
           #statSend.tsendFct.data[#statSend.tsendFct.dataOffset + 8] := #statSend.dataTelegram.ackMessageOffset.%B3;
           #statSend.tsendFct.data[#statSend.tsendFct.dataOffset + 9] := #statSend.dataTelegram.ackMessageOffset.%B2;
           #statSend.tsendFct.data[#statSend.tsendFct.dataOffset + 10] := #statSend.dataTelegram.ackMessageOffset.%B1;
           #statSend.tsendFct.data[#statSend.tsendFct.dataOffset + 11] := #statSend.dataTelegram.ackMessageOffset.%B0;

           #statSend.tsendFct.data[#statSend.tsendFct.dataOffset + 12] := #statSend.dataTelegram.actPackageLength.%B3;
           #statSend.tsendFct.data[#statSend.tsendFct.dataOffset + 13] := #statSend.dataTelegram.actPackageLength.%B2;
           #statSend.tsendFct.data[#statSend.tsendFct.dataOffset + 14] := #statSend.dataTelegram.actPackageLength.%B1;
           #statSend.tsendFct.data[#statSend.tsendFct.dataOffset + 15] := #statSend.dataTelegram.actPackageLength.%B0;

           #statSend.tsendFct.data[#statSend.tsendFct.dataOffset + 16] := #statSend.dataTelegram.totalMessageLength.%B3;
           #statSend.tsendFct.data[#statSend.tsendFct.dataOffset + 17] := #statSend.dataTelegram.totalMessageLength.%B2;
           #statSend.tsendFct.data[#statSend.tsendFct.dataOffset + 18] := #statSend.dataTelegram.totalMessageLength.%B1;
           #statSend.tsendFct.data[#statSend.tsendFct.dataOffset + 19] := #statSend.dataTelegram.totalMessageLength.%B0;

           //LCom V2
           IF (#diagnostics.statistics.activeLComVersion = #LCOM_HEADER_V2) THEN
             //Calculate offset in the tcp send buffer
             #statSend.tsendFct.dataOffset := #statSend.tsendFct.dataOffset + 20;
           ELSE
             //LCom V1
             //MessageOffset
             #statSend.tsendFct.data[#statSend.tsendFct.dataOffset + 4] := #statSend.dataTelegram.messageOffset.%B1;
             #statSend.tsendFct.data[#statSend.tsendFct.dataOffset + 5] := #statSend.dataTelegram.messageOffset.%B0;
             //AckMessageOffset
             #statSend.tsendFct.data[#statSend.tsendFct.dataOffset + 6] := #statSend.dataTelegram.ackMessageOffset.%B1;
             #statSend.tsendFct.data[#statSend.tsendFct.dataOffset + 7] := #statSend.dataTelegram.ackMessageOffset.%B0;
             //ActPackageLength
             #statSend.tsendFct.data[#statSend.tsendFct.dataOffset + 8] := #statSend.dataTelegram.actPackageLength.%B1;
             #statSend.tsendFct.data[#statSend.tsendFct.dataOffset + 9] := #statSend.dataTelegram.actPackageLength.%B0;
             //TotalMessageLength
             #statSend.tsendFct.data[#statSend.tsendFct.dataOffset + 10] := #statSend.dataTelegram.totalMessageLength.%B1;
             #statSend.tsendFct.data[#statSend.tsendFct.dataOffset + 11] := #statSend.dataTelegram.totalMessageLength.%B0;
             //Calculate offset in the tcp send buffer
             #statSend.tsendFct.dataOffset := #statSend.tsendFct.dataOffset + 12;
           END_IF;

           //Store expected acknowledge message offset and time
           #statSend.expectedAck.package1.offset := #statSend.dataTelegram.messageOffset + #statSend.dataTelegram.actPackageLength;
           //Start expe. message Timer 1
           #instExpectedAckPackage1(IN := TRUE,
                                    PT := #diagnostics.localConfig.sender.ackTimeout);

           #statSend.numberOfLComPackage := #statSend.numberOfLComPackage + 1;

           //Copy data from FB.sendBuffer
           #statRet := MOVE_BLK_VARIANT(SRC := #sendBuffer, COUNT := #statSend.dataTelegram.actPackageLength, SRC_INDEX := UDINT_TO_DINT(#statSend.userData.offset), DEST_INDEX := #statSend.tsendFct.dataOffset, DEST => #statSend.tsendFct.data);
           //Calculate offset in FB.sendBuffer
           #statSend.userData.offset := #statSend.userData.offset + #statSend.dataTelegram.actPackageLength;
           //Copy offset in telegram
           #statSend.dataTelegram.messageOffset := #statSend.userData.offset;
           //Calculate offset in the tcp send buffer
           #statSend.tsendFct.dataOffset := #statSend.tsendFct.dataOffset + UDINT_TO_UINT(#statSend.dataTelegram.actPackageLength);

           //All sent data is copied ?
           IF (#statSend.userData.offset = #statSend.dataTelegram.totalMessageLength) THEN
             //Yes
             #statState.comSender := #SEND_NO_DATA;
           ELSE
             ;//No --> Not all sent data has been copied
           END_IF;
         ELSIF (#statState.comSender = #CYCLE
           AND
           (NOT #diagnostics.localConfig.connection.useLComProtocol)) THEN
           //---------------------------------------------------------------------
           //Send telegram without LCom protocol
           //---------------------------------------------------------------------
           #statState.sender := #SEND_DATA;

           //Calculate rest data from the total message
           IF ((#statSend.dataTelegram.totalMessageLength - #statSend.userData.offset) > #MAX_DATA_BUFFER) THEN
             #statSend.tsendFct.dataOffset := #MAX_DATA_BUFFER;
           ELSE
             #statSend.tsendFct.dataOffset := UDINT_TO_UINT(#statSend.dataTelegram.totalMessageLength - #statSend.userData.offset);
           END_IF;

           //Copy data from FB.sendBuffer
           #statRet := MOVE_BLK_VARIANT(SRC := #sendBuffer, COUNT := #statSend.tsendFct.dataOffset, SRC_INDEX := UDINT_TO_DINT(#statSend.userData.offset), DEST_INDEX := 0, DEST => #statSend.tsendFct.data);
           //Calculate offset in tcp send buffer
           #statSend.userData.offset := #statSend.userData.offset + #statSend.tsendFct.dataOffset;
           //End: Send telegram without LCom protocol
         ELSE
           ;//Not in sending process 
         END_IF;//End: Send telegram
       END_IF;//End: Connected


       //---------------------------------------------------------------------
       //State machine sender configuration
       //---------------------------------------------------------------------
       CASE #statState.cfgSender OF

         #OPERATION:
           ;//Sender configuration successful exchange
         #STATE_WAIT:
           ;
         #STATE_INIT:

           #statCompare.sender.cycleTime := #configuration.sender.cycleTime;
           #statCompare.sender.ackTimeOut := #configuration.sender.ackTimeout;

           //LCom Version V1.0
           IF (#statActualLocalLComVersion = #LCOM_HEADER_V1) THEN

             //Check max. cycleTime
             IF (#configuration.sender.cycleTime > T#65535ms) THEN

               #statDiag.bufferIndex := #statDiag.bufferIndex + 1;
               #statDiag.buffer[#statDiag.bufferIndex].additionalValue4 := #configuration.sender.cycleTime;
               #statSend.configTelegramV1.cycleTime := 65535;

               #statDiag.buffer[#statDiag.bufferIndex].status := "LCOM_WARN_SEND_CYCLE_LIMITATION";
               #statDiag.buffer[#statDiag.bufferIndex].subFunctionErrorID := 16#0000;
               #statDiag.buffer[#statDiag.bufferIndex].additionalValue1 := 65535.0;
               #statDiag.buffer[#statDiag.bufferIndex].additionalValue2 := 0.0;
               #statDiag.buffer[#statDiag.bufferIndex].additionalValue3 := 0.0;
             ELSE
               #statSend.configTelegramV1.cycleTime := TIME_TO_UINT(#configuration.sender.cycleTime);
             END_IF;

             //Check max. ackTimeOut
             IF (#configuration.sender.ackTimeout > T#65535ms) THEN

               #statDiag.bufferIndex := #statDiag.bufferIndex + 1;
               #statDiag.buffer[#statDiag.bufferIndex].additionalValue4 := #configuration.sender.ackTimeout;
               #statSend.configTelegramV1.ackTimeOut := 65535;

               #statDiag.buffer[#statDiag.bufferIndex].status := "LCOM_WARN_ACK_TIMEOUT_LIMITATION";
               #statDiag.buffer[#statDiag.bufferIndex].subFunctionErrorID := 16#0000;
               #statDiag.buffer[#statDiag.bufferIndex].additionalValue1 := 65535.0;
               #statDiag.buffer[#statDiag.bufferIndex].additionalValue2 := 0.0;
               #statDiag.buffer[#statDiag.bufferIndex].additionalValue3 := 0.0;
             ELSE
               #statSend.configTelegramV1.ackTimeOut := TIME_TO_UINT(#configuration.sender.ackTimeout);
             END_IF;
           ELSE //LCom Version V2.0
             #statSend.configTelegramV2.cycleTime := #configuration.sender.cycleTime;
             #statSend.configTelegramV2.ackTimeOut := #configuration.sender.ackTimeout;
           END_IF;

           #statState.cfgSender := #SEND_CONFIG;

         #SEND_CONFIG:
           #statState.cfgSender := #STATE_WAIT;

           //LCom Version V1.0
           IF (#statActualLocalLComVersion = #LCOM_HEADER_V1) THEN
             #statSend.tsendFct.data[#statSend.tsendFct.dataOffset] := #statSend.configTelegramV1.LComVersion;
             #statSend.tsendFct.data[#statSend.tsendFct.dataOffset + 1] := 16#02;
             #statSend.tsendFct.data[#statSend.tsendFct.dataOffset + 2] := #statSend.configTelegramV1.comMode;//ComMode
             #statSend.tsendFct.data[#statSend.tsendFct.dataOffset + 3] := #statSend.configTelegramV1.slidingWindow;//SlidingWindow
             //cycleTime
             #statSend.tsendFct.data[#statSend.tsendFct.dataOffset + 4] := #statSend.configTelegramV1.cycleTime.%B1;
             #statSend.tsendFct.data[#statSend.tsendFct.dataOffset + 5] := #statSend.configTelegramV1.cycleTime.%B0;
             //ackTimeOut
             #statSend.tsendFct.data[#statSend.tsendFct.dataOffset + 6] := #statSend.configTelegramV1.ackTimeOut.%B1;
             #statSend.tsendFct.data[#statSend.tsendFct.dataOffset + 7] := #statSend.configTelegramV1.ackTimeOut.%B0;
             //lifeSignCycle
             #statSend.tsendFct.data[#statSend.tsendFct.dataOffset + 8] := #statSend.configTelegramV1.lifeSignCycle.%B1;
             #statSend.tsendFct.data[#statSend.tsendFct.dataOffset + 9] := #statSend.configTelegramV1.lifeSignCycle.%B0;
             //status
             #statSend.tsendFct.data[#statSend.tsendFct.dataOffset + 10] := #statSend.configTelegramV1.status;
             //sendModeSyncTime
             #statSend.tsendFct.data[#statSend.tsendFct.dataOffset + 11] := #statSend.configTelegramV1.sendModeSyncTime;
             //maxSendDataLength
             #statSend.tsendFct.data[#statSend.tsendFct.dataOffset + 12] := #statSend.configTelegramV1.maxSendDataLength.%B1;
             #statSend.tsendFct.data[#statSend.tsendFct.dataOffset + 13] := #statSend.configTelegramV1.maxSendDataLength.%B0;
             //maxReceiveDataLength
             #statSend.tsendFct.data[#statSend.tsendFct.dataOffset + 14] := #statSend.configTelegramV1.maxReceiveDataLength.%B1;
             #statSend.tsendFct.data[#statSend.tsendFct.dataOffset + 15] := #statSend.configTelegramV1.maxReceiveDataLength.%B0;

             #statSend.tsendFct.data[#statSend.tsendFct.dataOffset + 16] := #statSend.configTelegramV1.LComVersion;
             #statSend.tsendFct.data[#statSend.tsendFct.dataOffset + 17] := 16#02;
             #statSend.tsendFct.data[#statSend.tsendFct.dataOffset + 18] := #statSend.configTelegramV1.comMode;//ComMode
             #statSend.tsendFct.data[#statSend.tsendFct.dataOffset + 19] := #statSend.configTelegramV1.slidingWindow;//SlidingWindow
             //cycleTime
             #statSend.tsendFct.data[#statSend.tsendFct.dataOffset + 20] := #statSend.configTelegramV1.cycleTime.%B1;
             #statSend.tsendFct.data[#statSend.tsendFct.dataOffset + 21] := #statSend.configTelegramV1.cycleTime.%B0;
             //ackTimeOut
             #statSend.tsendFct.data[#statSend.tsendFct.dataOffset + 22] := #statSend.configTelegramV1.ackTimeOut.%B1;
             #statSend.tsendFct.data[#statSend.tsendFct.dataOffset + 23] := #statSend.configTelegramV1.ackTimeOut.%B0;
             //lifeSignCycle
             #statSend.tsendFct.data[#statSend.tsendFct.dataOffset + 24] := #statSend.configTelegramV1.lifeSignCycle.%B1;
             #statSend.tsendFct.data[#statSend.tsendFct.dataOffset + 25] := #statSend.configTelegramV1.lifeSignCycle.%B0;
             //status
             #statSend.tsendFct.data[#statSend.tsendFct.dataOffset + 26] := #statSend.configTelegramV1.status;
             //sendModeSyncTime
             #statSend.tsendFct.data[#statSend.tsendFct.dataOffset + 27] := #statSend.configTelegramV1.sendModeSyncTime;
             //maxSendDataLength
             #statSend.tsendFct.data[#statSend.tsendFct.dataOffset + 28] := #statSend.configTelegramV1.maxSendDataLength.%B1;
             #statSend.tsendFct.data[#statSend.tsendFct.dataOffset + 29] := #statSend.configTelegramV1.maxSendDataLength.%B0;
             //maxReceiveDataLength
             #statSend.tsendFct.data[#statSend.tsendFct.dataOffset + 30] := #statSend.configTelegramV1.maxReceiveDataLength.%B1;
             #statSend.tsendFct.data[#statSend.tsendFct.dataOffset + 31] := #statSend.configTelegramV1.maxReceiveDataLength.%B0;
             //calculate new offset
             #statSend.tsendFct.dataOffset := #statSend.tsendFct.dataOffset + 32;
             #statState.sender := #SEND_CONFIG;

             #diagnostics.localConfig.sender.cycleTime := UINT_TO_TIME(#statSend.configTelegramV1.cycleTime);
             #diagnostics.localConfig.sender.ackTimeout := UINT_TO_TIME(#statSend.configTelegramV1.ackTimeOut);
           ELSE
             //LCom Version V2.0
             #statSend.tsendFct.data[#statSend.tsendFct.dataOffset] := #statSend.configTelegramV2.LComVersion;
             #statSend.tsendFct.data[#statSend.tsendFct.dataOffset + 1] := 16#02;
             //status
             #statSend.tsendFct.data[#statSend.tsendFct.dataOffset + 2] := #statSend.configTelegramV2.status;
             //sendModeSyncTime
             #statSend.tsendFct.data[#statSend.tsendFct.dataOffset + 3] := #statSend.configTelegramV2.sendModeSyncTime;
             //lifeSignCycle
             #tempDWord := TIME_TO_DWORD(#statSend.configTelegramV2.lifeSignCycle);
             #statSend.tsendFct.data[#statSend.tsendFct.dataOffset + 4] := #tempDWord.%B3;
             #statSend.tsendFct.data[#statSend.tsendFct.dataOffset + 5] := #tempDWord.%B2;
             #statSend.tsendFct.data[#statSend.tsendFct.dataOffset + 6] := #tempDWord.%B1;
             #statSend.tsendFct.data[#statSend.tsendFct.dataOffset + 7] := #tempDWord.%B0;
             //cycleTime
             #tempDWord := TIME_TO_DWORD(#statSend.configTelegramV2.cycleTime);
             #statSend.tsendFct.data[#statSend.tsendFct.dataOffset + 8] := #tempDWord.%B3;
             #statSend.tsendFct.data[#statSend.tsendFct.dataOffset + 9] := #tempDWord.%B2;
             #statSend.tsendFct.data[#statSend.tsendFct.dataOffset + 10] := #tempDWord.%B1;
             #statSend.tsendFct.data[#statSend.tsendFct.dataOffset + 11] := #tempDWord.%B0;
             //ackTimeOut
             #tempDWord := TIME_TO_DWORD(#statSend.configTelegramV2.ackTimeOut);
             #statSend.tsendFct.data[#statSend.tsendFct.dataOffset + 12] := #tempDWord.%B3;
             #statSend.tsendFct.data[#statSend.tsendFct.dataOffset + 13] := #tempDWord.%B2;
             #statSend.tsendFct.data[#statSend.tsendFct.dataOffset + 14] := #tempDWord.%B1;
             #statSend.tsendFct.data[#statSend.tsendFct.dataOffset + 15] := #tempDWord.%B0;
             //maxSendDataLength
             #statSend.tsendFct.data[#statSend.tsendFct.dataOffset + 16] := #statSend.configTelegramV2.maxSendDataLength.%B3;
             #statSend.tsendFct.data[#statSend.tsendFct.dataOffset + 17] := #statSend.configTelegramV2.maxSendDataLength.%B2;
             #statSend.tsendFct.data[#statSend.tsendFct.dataOffset + 18] := #statSend.configTelegramV2.maxSendDataLength.%B1;
             #statSend.tsendFct.data[#statSend.tsendFct.dataOffset + 19] := #statSend.configTelegramV2.maxSendDataLength.%B0;
             //maxReceiveDataLength
             #statSend.tsendFct.data[#statSend.tsendFct.dataOffset + 20] := #statSend.configTelegramV2.maxReceiveDataLength.%B3;
             #statSend.tsendFct.data[#statSend.tsendFct.dataOffset + 21] := #statSend.configTelegramV2.maxReceiveDataLength.%B2;
             #statSend.tsendFct.data[#statSend.tsendFct.dataOffset + 22] := #statSend.configTelegramV2.maxReceiveDataLength.%B1;
             #statSend.tsendFct.data[#statSend.tsendFct.dataOffset + 23] := #statSend.configTelegramV2.maxReceiveDataLength.%B0;

             //calculate new offset
             #statSend.tsendFct.dataOffset := #statSend.tsendFct.dataOffset + 24;
             #statState.sender := #SEND_CONFIG;

             #diagnostics.localConfig.sender.cycleTime := #statSend.configTelegramV2.cycleTime;
             #diagnostics.localConfig.sender.ackTimeout := #statSend.configTelegramV2.ackTimeOut;

             IF #diagnostics.statistics.activeLComVersion = #LCOM_HEADER_V2 THEN
               #connected := TRUE;
               #diagnostics.statistics.LComProtocolUsed := TRUE;
               #diagnostics.statistics.activeLComVersion := #LCOM_HEADER_V2;
               #statState.cfgSender := #OPERATION;

               //Write diagnostics
               #statDiag.bufferIndex := #statDiag.bufferIndex + 1;
               #statDiag.buffer[#statDiag.bufferIndex].status := "LCOM_STATUS_LCOM_CONNECTED_V2";
               #statDiag.buffer[#statDiag.bufferIndex].subFunctionErrorID := 16#0000;
               #statDiag.buffer[#statDiag.bufferIndex].additionalValue1 := 0.0;
               #statDiag.buffer[#statDiag.bufferIndex].additionalValue2 := 0.0;
               #statDiag.buffer[#statDiag.bufferIndex].additionalValue3 := 0.0;
               #statDiag.buffer[#statDiag.bufferIndex].additionalValue4 := T#0ms;
             END_IF;
           END_IF;

           #statCompare.sender.cycleTime := #configuration.sender.cycleTime;
           #statCompare.sender.ackTimeOut := #configuration.sender.ackTimeout;

         #ERROR_STATE:
           ;
         ELSE
           ;// Statement section ELSE
       END_CASE;


       //No telegram 1,2,5 or 10 to  be sent, therefore check whether life sign tel. must be sent
       IF (#statState.sender = #STATE_INACTIVE
         AND
         (#diagnostics.localConfig.connection.lifeSignCycleTime <> T#0ms)
         AND
         #diagnostics.localConfig.connection.useLComProtocol)
       THEN
         #instLocalLifeSignCycleTimer(IN := TRUE,
                                      PT := #diagnostics.localConfig.connection.lifeSignCycleTime);

         IF (#instLocalLifeSignCycleTimer.Q)
         THEN

           //LCom Version V1.0
           IF (#statActualLocalLComVersion = #LCOM_HEADER_V1) THEN

             //LCom Version V1
             #statSend.tsendFct.data[#statSend.tsendFct.dataOffset] := #statSend.configTelegramV1.LComVersion;
             #statSend.tsendFct.data[#statSend.tsendFct.dataOffset + 1] := 16#03;
             #statSend.tsendFct.data[#statSend.tsendFct.dataOffset + 2] := #statSend.configTelegramV1.comMode;//ComMode
             #statSend.tsendFct.data[#statSend.tsendFct.dataOffset + 3] := #statSend.configTelegramV1.slidingWindow;//SlidingWindow
             //cycleTime
             #statSend.tsendFct.data[#statSend.tsendFct.dataOffset + 4] := #statSend.configTelegramV1.cycleTime.%B1;
             #statSend.tsendFct.data[#statSend.tsendFct.dataOffset + 5] := #statSend.configTelegramV1.cycleTime.%B0;
             //ackTimeOut
             #statSend.tsendFct.data[#statSend.tsendFct.dataOffset + 6] := #statSend.configTelegramV1.ackTimeOut.%B1;
             #statSend.tsendFct.data[#statSend.tsendFct.dataOffset + 7] := #statSend.configTelegramV1.ackTimeOut.%B0;
             //lifeSignCycle
             #statSend.tsendFct.data[#statSend.tsendFct.dataOffset + 8] := #statSend.configTelegramV1.lifeSignCycle.%B1;
             #statSend.tsendFct.data[#statSend.tsendFct.dataOffset + 9] := #statSend.configTelegramV1.lifeSignCycle.%B0;
             //status
             #statSend.tsendFct.data[#statSend.tsendFct.dataOffset + 10] := #statSend.configTelegramV1.status;
             //sendModeSyncTime
             #statSend.tsendFct.data[#statSend.tsendFct.dataOffset + 11] := #statSend.configTelegramV1.sendModeSyncTime;
             //maxSendDataLength
             #statSend.tsendFct.data[#statSend.tsendFct.dataOffset + 12] := #statSend.configTelegramV1.maxSendDataLength.%B1;
             #statSend.tsendFct.data[#statSend.tsendFct.dataOffset + 13] := #statSend.configTelegramV1.maxSendDataLength.%B0;
             //maxReceiveDataLength
             #statSend.tsendFct.data[#statSend.tsendFct.dataOffset + 14] := #statSend.configTelegramV1.maxReceiveDataLength.%B1;
             #statSend.tsendFct.data[#statSend.tsendFct.dataOffset + 15] := #statSend.configTelegramV1.maxReceiveDataLength.%B0;
             //calculate new offset
             #statSend.tsendFct.dataOffset := 16;
           ELSE
             #statSend.tsendFct.data[#statSend.tsendFct.dataOffset] := #statSend.configTelegramV2.LComVersion;
             #statSend.tsendFct.data[#statSend.tsendFct.dataOffset + 1] := 16#03;
             //status
             #statSend.tsendFct.data[#statSend.tsendFct.dataOffset + 2] := #statSend.configTelegramV2.status;
             //sendModeSyncTime
             #statSend.tsendFct.data[#statSend.tsendFct.dataOffset + 3] := #statSend.configTelegramV2.sendModeSyncTime;
             //lifeSignCycle
             #tempDWord := TIME_TO_DWORD(#statSend.configTelegramV2.lifeSignCycle);
             #statSend.tsendFct.data[#statSend.tsendFct.dataOffset + 4] := #tempDWord.%B3;
             #statSend.tsendFct.data[#statSend.tsendFct.dataOffset + 5] := #tempDWord.%B2;
             #statSend.tsendFct.data[#statSend.tsendFct.dataOffset + 6] := #tempDWord.%B1;
             #statSend.tsendFct.data[#statSend.tsendFct.dataOffset + 7] := #tempDWord.%B0;
             //cycleTime
             #tempDWord := TIME_TO_DWORD(#statSend.configTelegramV2.cycleTime);
             #statSend.tsendFct.data[#statSend.tsendFct.dataOffset + 8] := #tempDWord.%B3;
             #statSend.tsendFct.data[#statSend.tsendFct.dataOffset + 9] := #tempDWord.%B2;
             #statSend.tsendFct.data[#statSend.tsendFct.dataOffset + 10] := #tempDWord.%B1;
             #statSend.tsendFct.data[#statSend.tsendFct.dataOffset + 11] := #tempDWord.%B0;
             //ackTimeOut
             #tempDWord := TIME_TO_DWORD(#statSend.configTelegramV2.ackTimeOut);
             #statSend.tsendFct.data[#statSend.tsendFct.dataOffset + 12] := #tempDWord.%B3;
             #statSend.tsendFct.data[#statSend.tsendFct.dataOffset + 13] := #tempDWord.%B2;
             #statSend.tsendFct.data[#statSend.tsendFct.dataOffset + 14] := #tempDWord.%B1;
             #statSend.tsendFct.data[#statSend.tsendFct.dataOffset + 15] := #tempDWord.%B0;
             //maxSendDataLength
             #statSend.tsendFct.data[#statSend.tsendFct.dataOffset + 16] := #statSend.configTelegramV2.maxSendDataLength.%B3;
             #statSend.tsendFct.data[#statSend.tsendFct.dataOffset + 17] := #statSend.configTelegramV2.maxSendDataLength.%B2;
             #statSend.tsendFct.data[#statSend.tsendFct.dataOffset + 18] := #statSend.configTelegramV2.maxSendDataLength.%B1;
             #statSend.tsendFct.data[#statSend.tsendFct.dataOffset + 19] := #statSend.configTelegramV2.maxSendDataLength.%B0;
             //maxReceiveDataLength
             #statSend.tsendFct.data[#statSend.tsendFct.dataOffset + 20] := #statSend.configTelegramV2.maxReceiveDataLength.%B3;
             #statSend.tsendFct.data[#statSend.tsendFct.dataOffset + 21] := #statSend.configTelegramV2.maxReceiveDataLength.%B2;
             #statSend.tsendFct.data[#statSend.tsendFct.dataOffset + 22] := #statSend.configTelegramV2.maxReceiveDataLength.%B1;
             #statSend.tsendFct.data[#statSend.tsendFct.dataOffset + 23] := #statSend.configTelegramV2.maxReceiveDataLength.%B0;
             //calculate new offset
             #statSend.tsendFct.dataOffset := 24;
           END_IF;
           #statSend.tsendFct.enable := TRUE;

           #instLocalLifeSignCycleTimer(IN := FALSE,
                                        PT := #diagnostics.localConfig.connection.lifeSignCycleTime);
         ELSE
           ;//Telegram 3 don´t need be send

         END_IF;
       ELSIF (NOT #diagnostics.localConfig.connection.useLComProtocol //without LCom Protocol
         AND #statState.sender = #STATE_INACTIVE) THEN
         #statSend.tsendFct.enable := FALSE;
       ELSE
         #statSend.tsendFct.enable := TRUE;

         #instLocalLifeSignCycleTimer(IN := FALSE,
                                      PT := #diagnostics.localConfig.connection.lifeSignCycleTime);
       END_IF;

       #instTSEND(REQ := #statSend.tsendFct.enable,
                  LEN := #statSend.tsendFct.dataOffset,
                  ID := #statTconPar.ID,
                  DATA := #statSend.tsendFct.data,
                  STATUS => #statSend.tsendFct.status);

       //16#80C4=Temporary communication error
       IF (#statSend.tsendFct.status = 16#80C4) THEN

         #instSendErrorTimer(IN := TRUE,
                             PT := #MAX_TRIAL_TIME);

         //#MAX_TRIAL_TIME is expired
         IF #instSendErrorTimer.Q THEN
           //Write diagnostics
           #statDiag.bufferIndex := #statDiag.bufferIndex + 1;
           #statDiag.buffer[#statDiag.bufferIndex].status := "LCOM_ERR_SEND";
           #statDiag.buffer[#statDiag.bufferIndex].subFunctionErrorID := #statSend.tsendFct.status;
           #statDiag.buffer[#statDiag.bufferIndex].additionalValue1 := 0.0;
           #statDiag.buffer[#statDiag.bufferIndex].additionalValue2 := #statSend.tsendFct.dataOffset;
           #statDiag.buffer[#statDiag.bufferIndex].additionalValue3 := 0.0;
           #statDiag.buffer[#statDiag.bufferIndex].additionalValue4 := T#0ms;
           #statState.connection := #CLOSE_CONNECTION;
           GOTO diag;
         END_IF;
       ELSIF (#statSend.tsendFct.status >= 16#8085) THEN
         //#WARN_SEND
         #statDiag.bufferIndex := #statDiag.bufferIndex + 1;
         #statDiag.buffer[#statDiag.bufferIndex].status := "LCOM_ERR_SEND";
         #statDiag.buffer[#statDiag.bufferIndex].subFunctionErrorID := #statSend.tsendFct.status;
         #statDiag.buffer[#statDiag.bufferIndex].additionalValue1 := 0.0;
         #statDiag.buffer[#statDiag.bufferIndex].additionalValue2 := #statSend.tsendFct.dataOffset;
         #statDiag.buffer[#statDiag.bufferIndex].additionalValue3 := 0.0;
         #statDiag.buffer[#statDiag.bufferIndex].additionalValue4 := T#0ms;

         #statState.connection := #CLOSE_CONNECTION;
         GOTO diag;
       END_IF;

     #STATE_INACTIVE_PREPARE:

       #statState.connection := #STATE_INACTIVE;
       #status := "LCOM_STATUS_NO_CALL";
       #statFallingEdgeEnable := FALSE;
       #statOldEnable := FALSE;
       #busy := FALSE;

     #STATE_INIT:
       //Reset FB Outputs
       #connected := FALSE;
       #sending := FALSE;
       #error := FALSE;

       //Diagnostics purpose
       //connection
       #diagnostics.localConfig.connection.connectionID := #configuration.connection.connectionID;
       #diagnostics.localConfig.connection.interfaceID := #configuration.connection.interfaceID;
       #diagnostics.localConfig.connection.comService := #configuration.connection.comService;
       #diagnostics.localConfig.connection.isClient := #configuration.connection.isClient;
       #diagnostics.localConfig.connection.localPort := #configuration.connection.localPort;
       #diagnostics.localConfig.connection.partnerPort := #configuration.connection.partnerPort;
       #diagnostics.localConfig.connection.partnerIP := #configuration.connection.partnerIP;
       #diagnostics.localConfig.connection.acceptUnknownPartner := #configuration.connection.acceptUnknownPartner;
       #statActualLocalLComVersion := #LCOM_HEADER_V2;
       #diagnostics.localConfig.connection.lifeSignCycleTime := #configuration.connection.lifeSignCycleTime;
       //Sender
       #diagnostics.localConfig.sender.cycleTime := #configuration.sender.cycleTime;
       #diagnostics.localConfig.sender.ackTimeout := #configuration.sender.ackTimeout;
       //TimeSync
       #diagnostics.localConfig.timeSync.usePartnerTimestamps := #configuration.timeSync.usePartnerTimestamps;
       #diagnostics.localConfig.timeSync.sendMode := #configuration.timeSync.sendMode;
       #diagnostics.localConfig.timeSync.cycleTime := #configuration.timeSync.cycleTime;
       #diagnostics.localConfig.timeSync.sendAtTimeOfDay := #configuration.timeSync.sendAtTimeOfDay;
       //Statistics
       #diagnostics.statistics.avgCallCycle := 0.0;
       #diagnostics.statistics.avgReceiveMsgCycle := 0.0;
       #diagnostics.statistics.maxReceiveMsgCycle := T#0ms;
       #diagnostics.statistics.LComProtocolUsed := FALSE;
       #diagnostics.statistics.activeLComVersion := 0;
       #diagnostics.statistics.avgMsgSendingTime := 0.0;
       #diagnostics.statistics.maxMsgSendingTime := T#0ms;
       #diagnostics.statistics.avgMsgReceivingTime := 0.0;
       #diagnostics.statistics.maxMsgReceivingTime := T#0ms;
       #diagnostics.statistics.numberOfSentMessages := 0;
       #diagnostics.statistics.numberOfReceivedMessages := 0;
       #diagnostics.statistics.totalAckTimeouts := 0;
       #diagnostics.statistics.totalSendCycleViolations := 0;
       #diagnostics.statistics.totalReceiveCycleViolations := 0;
       #diagnostics.statistics.totalReconnects := 0;

       #statConnectAttempts := 0;

       //Check hardware identifier of the local interface
       IF ((#diagnostics.localConfig.connection.interfaceID >= 0) //(0...65535)
         AND
         (#diagnostics.localConfig.connection.interfaceID <= 65535))
       THEN
         //Hardware identifier of the local interface --> OK
         #statTconPar.InterfaceId := #diagnostics.localConfig.connection.interfaceID;
       ELSE
         //Hardware identifier of the local interface --> NOT OK
         #statDiag.bufferIndex := #statDiag.bufferIndex + 1;
         #statDiag.buffer[#statDiag.bufferIndex].status := "LCOM_ERR_INTERFACE_ID";
         #statDiag.buffer[#statDiag.bufferIndex].subFunctionErrorID := 16#0000;
         #statDiag.buffer[#statDiag.bufferIndex].additionalValue1 := UINT_TO_REAL(#diagnostics.localConfig.connection.interfaceID);//value from user
         #statDiag.buffer[#statDiag.bufferIndex].additionalValue2 := 0.0;
         #statDiag.buffer[#statDiag.bufferIndex].additionalValue3 := 0.0;
         #statDiag.buffer[#statDiag.bufferIndex].additionalValue4 := T#0ms;

         #statState.connection := #ERROR_STATE;
         GOTO diag;
       END_IF;

       //Read the IP address
       #instRDREC(REQ := TRUE,
                  ID := #configuration.connection.interfaceID,
                  INDEX := 16#8080,
                  MLEN := 0,
                  RECORD := #statSend.tsendFct.data);

       //1st call from RDREC, to get the IP address
       IF #instRDREC.STATUS = 16#00700100 THEN
           ;//don´t change the #status = "LCOM_STATUS_FIRST_CALL"
       ELSE
           //change status, that 1st call is just one time occur 
           #status := "LCOM_STATUS_INTERMEDIATE_CALL";
       END_IF;

       IF (#instRDREC.VALID = TRUE) THEN
         //New data received and data is valid
         #diagnostics.localConfig.connection.localIP.ADDR[1] := #statSend.tsendFct.data[28];
         #diagnostics.localConfig.connection.localIP.ADDR[2] := #statSend.tsendFct.data[29];
         #diagnostics.localConfig.connection.localIP.ADDR[3] := #statSend.tsendFct.data[30];
         #diagnostics.localConfig.connection.localIP.ADDR[4] := #statSend.tsendFct.data[31];
       ELSIF (#instRDREC.ERROR = TRUE) THEN
         //An error occurred during the reading process
         #diagnostics.localConfig.connection.localIP.ADDR[1] := 16#00;
         #diagnostics.localConfig.connection.localIP.ADDR[2] := 16#00;
         #diagnostics.localConfig.connection.localIP.ADDR[3] := 16#00;
         #diagnostics.localConfig.connection.localIP.ADDR[4] := 16#00;
       ELSE
         RETURN;//The reading process is not complete yet
       END_IF;

       //Local port number
       #statTconPar.LocalPort := #diagnostics.localConfig.connection.localPort;

       //Check if send buffer is a VARIANT pointer to array of byte
       IF ((TypeOfElements(#sendBuffer) = TypeOf(#statSend.tsendFct.data[0]))
         AND
         (IS_ARRAY(#sendBuffer))) THEN
         ;//Is VARIANT pointer to array of byte
       ELSE
         //Write diagnostics
         #statDiag.bufferIndex := #statDiag.bufferIndex + 1;
         #statDiag.buffer[#statDiag.bufferIndex].status := "LCOM_ERR_SEND_DATA_TYPE";
         #statDiag.buffer[#statDiag.bufferIndex].subFunctionErrorID := 16#0000;
         #statDiag.buffer[#statDiag.bufferIndex].additionalValue1 := 0.0;
         #statDiag.buffer[#statDiag.bufferIndex].additionalValue2 := 0.0;
         #statDiag.buffer[#statDiag.bufferIndex].additionalValue3 := 0.0;
         #statDiag.buffer[#statDiag.bufferIndex].additionalValue4 := T#0ms;

         #statState.connection := #ERROR_STATE;
         GOTO diag;
       END_IF;

       //Check if receive buffer is a VARIANT pointer to array of byte
       IF ((TypeOfElements(#receiveBuffer) = TypeOf(#statReceive.trcvFct.data[0]))
         AND
         (IS_ARRAY(#receiveBuffer))) THEN
         ;//Is VARIANT pointer to array of byte
       ELSE
         //Write diagnostics
         #statDiag.bufferIndex := #statDiag.bufferIndex + 1;
         #statDiag.buffer[#statDiag.bufferIndex].status := "LCOM_ERR_RECEIVE_DATA_TYPE";
         #statDiag.buffer[#statDiag.bufferIndex].subFunctionErrorID := 16#0000;
         #statDiag.buffer[#statDiag.bufferIndex].additionalValue1 := 0.0;
         #statDiag.buffer[#statDiag.bufferIndex].additionalValue2 := 0.0;
         #statDiag.buffer[#statDiag.bufferIndex].additionalValue3 := 0.0;
         #statDiag.buffer[#statDiag.bufferIndex].additionalValue4 := T#0ms;

         #statState.connection := #ERROR_STATE;
         GOTO diag;
       END_IF;

       //Get size of user send buffer and user receive buffer in bytes
       #diagnostics.localConfig.sizeOfSendBuffer := CountOfElements(#sendBuffer);
       #diagnostics.localConfig.sizeOfReceiveBuffer := CountOfElements(#receiveBuffer);

       //Check communication service: 0:UDP, 1:TCP, 2:LCOM
       IF (#diagnostics.localConfig.connection.comService = 16#01) THEN
         //Communication service --> transport protocol TCP
         #statTconPar.ConnectionType := 16#0B;
         #diagnostics.localConfig.connection.useLComProtocol := FALSE;
       ELSIF (#diagnostics.localConfig.connection.comService = 16#02) THEN
         //Communication service --> transport protocol TCP and LCom protocol
         #statTconPar.ConnectionType := 16#0B;
         #diagnostics.localConfig.connection.useLComProtocol := TRUE;
       ELSE
         //Communication service --> NOT OK
         //Write diagnostics
         #statDiag.bufferIndex := #statDiag.bufferIndex + 1;
         #statDiag.buffer[#statDiag.bufferIndex].status := "LCOM_ERR_COM_SERVICE";
         #statDiag.buffer[#statDiag.bufferIndex].subFunctionErrorID := 16#0000;
         #statDiag.buffer[#statDiag.bufferIndex].additionalValue1 := #diagnostics.localConfig.connection.comService;//value from operator
         #statDiag.buffer[#statDiag.bufferIndex].additionalValue2 := 0.0;
         #statDiag.buffer[#statDiag.bufferIndex].additionalValue3 := 0.0;
         #statDiag.buffer[#statDiag.bufferIndex].additionalValue4 := T#0ms;

         #statState.connection := #ERROR_STATE;
         GOTO diag;
       END_IF;

       //Check unique connection identifier (16#0001...16#0FFF)
       IF ((#diagnostics.localConfig.connection.connectionID > 0)
         AND
         (#diagnostics.localConfig.connection.connectionID <= 4095))
       THEN
         //Connection identifier -->OK
         #statTconPar.ID := #diagnostics.localConfig.connection.connectionID;
       ELSE
         //Connection identifier --> NOT OK
         //Write diagnostics
         #statDiag.bufferIndex := #statDiag.bufferIndex + 1;
         #statDiag.buffer[#statDiag.bufferIndex].status := "LCOM_ERR_CONNECTION_ID";
         #statDiag.buffer[#statDiag.bufferIndex].subFunctionErrorID := 16#0000;
         #statDiag.buffer[#statDiag.bufferIndex].additionalValue1 := WORD_TO_UDINT(#diagnostics.localConfig.connection.connectionID);//value from user
         #statDiag.buffer[#statDiag.bufferIndex].additionalValue2 := 0.0;
         #statDiag.buffer[#statDiag.bufferIndex].additionalValue3 := 0.0;
         #statDiag.buffer[#statDiag.bufferIndex].additionalValue4 := T#0ms;

         #statState.connection := #ERROR_STATE;
         GOTO diag;
       END_IF;

       //If client
       IF (#diagnostics.localConfig.connection.isClient) THEN
         //Partner port and remote address is not checked here
         //The TCON will rise an error and return value, when the parameters (partnerPort or partnerIP) are wrong
         #statTconPar.RemotePort := #diagnostics.localConfig.connection.partnerPort;
         #statTconPar.RemoteAddress := #diagnostics.localConfig.connection.partnerIP;
       ELSE
         //If server
         //Accept requests from all partners or only specified partner is allowed
         IF (#diagnostics.localConfig.connection.acceptUnknownPartner) THEN
           //Accept requests from all partners
           #statTconPar.RemoteAddress.ADDR[1] := 0;
           #statTconPar.RemoteAddress.ADDR[2] := 0;
           #statTconPar.RemoteAddress.ADDR[3] := 0;
           #statTconPar.RemoteAddress.ADDR[4] := 0;
           #statTconPar.RemotePort := 0;
         ELSE
           //Only specified partner is allowed
           #statTconPar.RemoteAddress := #diagnostics.localConfig.connection.partnerIP;
           #statTconPar.RemotePort := #diagnostics.localConfig.connection.partnerPort;
         END_IF;
       END_IF;

       //Check cycleTime
       IF ((#diagnostics.localConfig.sender.cycleTime >= T#0ms)
         AND
         (#diagnostics.localConfig.sender.cycleTime <= T#+24d20h31m23s647ms))
       THEN
         ;//CycleTime --> OK
       ELSE
         //CycleTime --> NOT OK
         #statDiag.bufferIndex := #statDiag.bufferIndex + 1;
         #statDiag.buffer[#statDiag.bufferIndex].status := "LCOM_ERR_SEND_CYCLE_TIME";
         #statDiag.buffer[#statDiag.bufferIndex].subFunctionErrorID := 16#0000;
         #statDiag.buffer[#statDiag.bufferIndex].additionalValue1 := 0.0;
         #statDiag.buffer[#statDiag.bufferIndex].additionalValue2 := 0.0;
         #statDiag.buffer[#statDiag.bufferIndex].additionalValue3 := 0.0;
         #statDiag.buffer[#statDiag.bufferIndex].additionalValue4 := #diagnostics.localConfig.sender.cycleTime;//value from operator

         #statState.connection := #ERROR_STATE;
         GOTO diag;
       END_IF;

       //With LCom header
       IF (#diagnostics.localConfig.connection.useLComProtocol) THEN

         //Check lifeSignCycleTime
         IF ((#diagnostics.localConfig.connection.lifeSignCycleTime > T#0ms) //(1ms...T#+24d20h31m23s647ms)
           AND
           (#diagnostics.localConfig.connection.lifeSignCycleTime <= T#+24d20h31m23s647ms))
         THEN
           ;//lifeSignCycleTime--> OK
         ELSE
           //LifeSignCycle --> NOT OK
           #statDiag.bufferIndex := #statDiag.bufferIndex + 1;
           #statDiag.buffer[#statDiag.bufferIndex].status := "LCOM_ERR_LIFE_SIGN_CYCLE";
           #statDiag.buffer[#statDiag.bufferIndex].subFunctionErrorID := 16#0000;
           #statDiag.buffer[#statDiag.bufferIndex].additionalValue1 := 0.0;
           #statDiag.buffer[#statDiag.bufferIndex].additionalValue2 := 0.0;
           #statDiag.buffer[#statDiag.bufferIndex].additionalValue3 := 0.0;
           #statDiag.buffer[#statDiag.bufferIndex].additionalValue4 := #diagnostics.localConfig.connection.lifeSignCycleTime;//value from operator

           #statState.connection := #ERROR_STATE;
           GOTO diag;
         END_IF;

         //Check ackTimeOut
         IF ((#diagnostics.localConfig.sender.ackTimeout > T#0ms)
           AND
           (#diagnostics.localConfig.sender.ackTimeout <= T#+24d20h31m23s647ms))
         THEN
           ;//AckTimeOut --> OK
         ELSE
           //AckTimeOut --> NOT OK
           #statDiag.bufferIndex := #statDiag.bufferIndex + 1;
           #statDiag.buffer[#statDiag.bufferIndex].status := "LCOM_ERR_ACK_TIMEOUT";
           #statDiag.buffer[#statDiag.bufferIndex].subFunctionErrorID := 16#0000;
           #statDiag.buffer[#statDiag.bufferIndex].additionalValue1 := 0.0;
           #statDiag.buffer[#statDiag.bufferIndex].additionalValue2 := 0.0;
           #statDiag.buffer[#statDiag.bufferIndex].additionalValue3 := 0.0;
           #statDiag.buffer[#statDiag.bufferIndex].additionalValue4 := #diagnostics.localConfig.sender.ackTimeout;//value from operator

           #statState.connection := #ERROR_STATE;
           GOTO diag;
         END_IF;

         //Check timeSync
         IF (NOT #diagnostics.localConfig.timeSync.usePartnerTimestamps) THEN

           IF ((#diagnostics.localConfig.timeSync.sendMode >= 0)//(0...2)
             AND
             (#diagnostics.localConfig.timeSync.sendMode <= 2))
           THEN
             CASE (#diagnostics.localConfig.timeSync.sendMode) OF

               1: //TimeSync.cycleTime
                 IF ((#diagnostics.localConfig.timeSync.cycleTime > T#0ms) //(1ms...T#+24d20h31m23s647ms)
                   AND
                   (#diagnostics.localConfig.timeSync.cycleTime <= T#+24d20h31m23s647ms))
                 THEN
                   ;//CycleTime --> OK
                 ELSE
                   //CycleTime --> Not OK
                   #statDiag.bufferIndex := #statDiag.bufferIndex + 1;
                   #statDiag.buffer[#statDiag.bufferIndex].status := "LCOM_ERR_TIME_CYCLE_TIME";
                   #statDiag.buffer[#statDiag.bufferIndex].subFunctionErrorID := 16#0000;
                   #statDiag.buffer[#statDiag.bufferIndex].additionalValue1 := 0.0;
                   #statDiag.buffer[#statDiag.bufferIndex].additionalValue2 := 0.0;
                   #statDiag.buffer[#statDiag.bufferIndex].additionalValue3 := 0.0;
                   #statDiag.buffer[#statDiag.bufferIndex].additionalValue4 := #diagnostics.localConfig.timeSync.cycleTime;//value from user

                   #statState.connection := #ERROR_STATE;
                   GOTO diag;

                 END_IF;
               2://TimeSync.sendAtTimeOfDay
                 IF ((#diagnostics.localConfig.timeSync.sendAtTimeOfDay >= TOD#00:00:00.000) //(TOD#00:00:00.000...TOD#23:59:59.999)
                   AND
                   #diagnostics.localConfig.timeSync.sendAtTimeOfDay <= TOD#23:59:59.999)
                 THEN
                   ;//SendAtTimeOfDay --> OK
                 ELSE
                   //SendAtTimeOfDay --> NOT OK
                   #statDiag.bufferIndex := #statDiag.bufferIndex + 1;
                   #statDiag.buffer[#statDiag.bufferIndex].status := "LCOM_ERR_TIME_OF_DAY";
                   #statDiag.buffer[#statDiag.bufferIndex].subFunctionErrorID := 16#0000;
                   #statDiag.buffer[#statDiag.bufferIndex].additionalValue1 := 0.0;
                   #statDiag.buffer[#statDiag.bufferIndex].additionalValue2 := 0.0;
                   #statDiag.buffer[#statDiag.bufferIndex].additionalValue3 := 0.0;
                   #statDiag.buffer[#statDiag.bufferIndex].additionalValue4 := T#0ms;

                   #statState.connection := #ERROR_STATE;
                   GOTO diag;
                 END_IF;
               ELSE
                 ;
             END_CASE;
           ELSE
             //SendMode --> NOT OK
             #statDiag.bufferIndex := #statDiag.bufferIndex + 1;
             #statDiag.buffer[#statDiag.bufferIndex].status := "LCOM_ERR_TIME_SYNC_MODE";
             #statDiag.buffer[#statDiag.bufferIndex].subFunctionErrorID := 16#0000;
             #statDiag.buffer[#statDiag.bufferIndex].additionalValue1 := #diagnostics.localConfig.timeSync.sendMode;
             #statDiag.buffer[#statDiag.bufferIndex].additionalValue2 := 0.0;
             #statDiag.buffer[#statDiag.bufferIndex].additionalValue3 := 0.0;
             #statDiag.buffer[#statDiag.bufferIndex].additionalValue4 := T#0ms;

             #statState.connection := #ERROR_STATE;
             GOTO diag;
           END_IF;
         ELSE
           //usePartnerTimeStamp

           //Is sendMode inactive ?
           IF #diagnostics.localConfig.timeSync.sendMode = 0 THEN
             ;// Yes
           ELSE
             //SendMode --> NOT OK
             #statDiag.bufferIndex := #statDiag.bufferIndex + 1;
             #statDiag.buffer[#statDiag.bufferIndex].status := "LCOM_ERR_TIME_SYNC_MODE";
             #statDiag.buffer[#statDiag.bufferIndex].subFunctionErrorID := 16#0000;
             #statDiag.buffer[#statDiag.bufferIndex].additionalValue1 := #diagnostics.localConfig.timeSync.sendMode;
             #statDiag.buffer[#statDiag.bufferIndex].additionalValue2 := 0.0;
             #statDiag.buffer[#statDiag.bufferIndex].additionalValue3 := 0.0;
             #statDiag.buffer[#statDiag.bufferIndex].additionalValue4 := T#0ms;

             #statState.connection := #ERROR_STATE;
             GOTO diag;
           END_IF;

         END_IF;
       ELSE
         ;//No LCom Protocol is used
       END_IF;

       #instTCON(REQ := FALSE,
                 ID := #statTconPar.ID,
                 CONNECT := #statTconPar);

       #instTSEND(REQ := FALSE,
                  ID := #statTconPar.ID,
                  DATA := #statSend.tsendFct.data);

       #instTRCV(EN_R := FALSE,
                 ID := #statTconPar.ID,
                 DATA := #statReceive.trcvFct.data);

       #instTDISCON(REQ := FALSE,
                    ID := #statTconPar.ID);

       //Passive (server), active connection establishment (client)
       IF (#diagnostics.localConfig.connection.isClient) THEN
         #statState.connection := #OPEN_CLIENT;
         #statTconPar.ActiveEstablished := TRUE;
       ELSE
         #statState.connection := #OPEN_SERVER;
         #statTconPar.ActiveEstablished := FALSE;
       END_IF;

     #OPEN_CLIENT, #OPEN_SERVER:

       #instTCON.STATUS := 16#0000;

       #instTCON(REQ := TRUE,
                 CONNECT := #statTconPar,
                 ID := #diagnostics.localConfig.connection.connectionID);

       // Error occurred
       IF (#instTCON.ERROR) THEN

           //Local port is being used by the system
           IF (#instTCON.STATUS = 16#80A2 OR #statTconPar.LocalPort=16#0) THEN

           #statDiag.bufferIndex := #statDiag.bufferIndex + 1;
           #statDiag.buffer[#statDiag.bufferIndex].status := "LCOM_ERR_LOCAL_PORT";
           #statDiag.buffer[#statDiag.bufferIndex].subFunctionErrorID := #instTCON.STATUS;
           #statDiag.buffer[#statDiag.bufferIndex].additionalValue1 := #statTconPar.LocalPort;
           #statDiag.buffer[#statDiag.bufferIndex].additionalValue2 := 0.0;
           #statDiag.buffer[#statDiag.bufferIndex].additionalValue3 := 0.0;
           #statDiag.buffer[#statDiag.bufferIndex].additionalValue4 := T#0ms;

           #statState.connection := #ERROR_STATE;
           GOTO diag;
         ELSIF (#instTCON.STATUS = 16#80B7 OR #instTCON.STATUS = 16#80A4) THEN
           //IP address of the remote partner is invalid
           #statDiag.bufferIndex := #statDiag.bufferIndex + 1;
           #statDiag.buffer[#statDiag.bufferIndex].status := "LCOM_ERR_PARTNER_IP";
           #statDiag.buffer[#statDiag.bufferIndex].subFunctionErrorID := #instTCON.STATUS;
           #statDiag.buffer[#statDiag.bufferIndex].additionalValue1 := 0.0;
           #statDiag.buffer[#statDiag.bufferIndex].additionalValue2 := 0.0;
           #statDiag.buffer[#statDiag.bufferIndex].additionalValue3 := 0.0;
           #statDiag.buffer[#statDiag.bufferIndex].additionalValue4 := T#0ms;

           #statState.connection := #ERROR_STATE;
           GOTO diag;
         ELSIF (#instTCON.STATUS = 16#809B) THEN
           //The local_device_id in the connection description does not match the CPU
           #statDiag.bufferIndex := #statDiag.bufferIndex + 1;
           #statDiag.buffer[#statDiag.bufferIndex].status := "LCOM_ERR_INTERFACE_ID";
           #statDiag.buffer[#statDiag.bufferIndex].subFunctionErrorID := #instTCON.STATUS;
           #statDiag.buffer[#statDiag.bufferIndex].additionalValue1 := UINT_TO_REAL(#diagnostics.localConfig.connection.interfaceID);//value from user
           #statDiag.buffer[#statDiag.bufferIndex].additionalValue2 := 0.0;
           #statDiag.buffer[#statDiag.bufferIndex].additionalValue3 := 0.0;
           #statDiag.buffer[#statDiag.bufferIndex].additionalValue4 := T#0ms;

           #statState.connection := #ERROR_STATE;
           GOTO diag;
         ELSE
           IF (#statState.connection = #OPEN_CLIENT) THEN

             #statDiag.bufferIndex := #statDiag.bufferIndex + 1;
             #statDiag.buffer[#statDiag.bufferIndex].status := "LCOM_ERR_OPEN_CLIENT";
             #statDiag.buffer[#statDiag.bufferIndex].subFunctionErrorID := #instTCON.STATUS;
             #statDiag.buffer[#statDiag.bufferIndex].additionalValue1 := 0.0;
             #statDiag.buffer[#statDiag.bufferIndex].additionalValue2 := 0.0;
             #statDiag.buffer[#statDiag.bufferIndex].additionalValue3 := 0.0;
             #statDiag.buffer[#statDiag.bufferIndex].additionalValue4 := T#0ms;

             //Try reconnection after a wait time
             #statIterator := 0;
             #statState.connection := #STATE_WAIT;
           ELSE
             #statDiag.bufferIndex := #statDiag.bufferIndex + 1;
             #statDiag.buffer[#statDiag.bufferIndex].status := "LCOM_ERR_OPEN_SERVER";
             #statDiag.buffer[#statDiag.bufferIndex].subFunctionErrorID := #instTCON.STATUS;
             #statDiag.buffer[#statDiag.bufferIndex].additionalValue1 := #statTconPar.LocalPort;
             #statDiag.buffer[#statDiag.bufferIndex].additionalValue2 := 0.0;
             #statDiag.buffer[#statDiag.bufferIndex].additionalValue3 := 0.0;
             #statDiag.buffer[#statDiag.bufferIndex].additionalValue4 := T#0ms;

